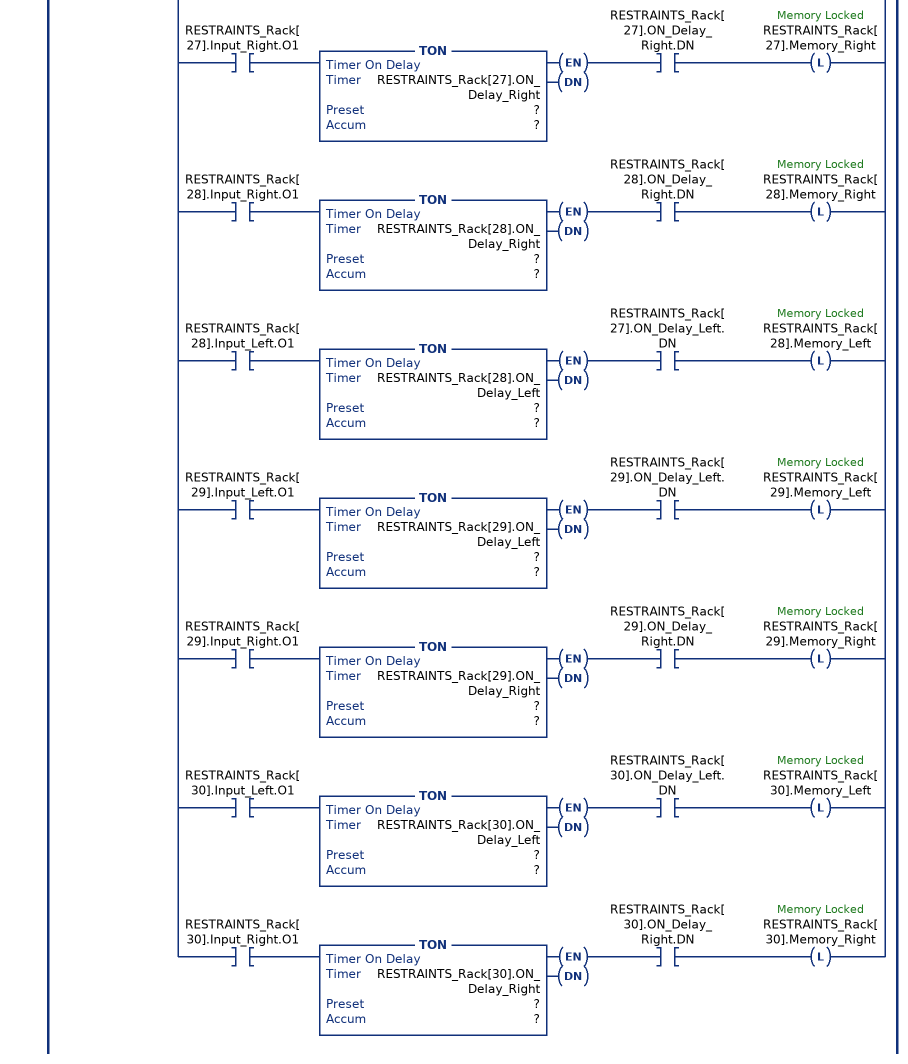
   14: XIC(Restraints_Cycle.Step_22)[XIC(RESTRAINTS_Rack[17].Input_Left.O1) TON(RESTRAINTS_Rack[17].ON_Delay_Left,?,?) XIC(RESTRAINTS_Rack[17].ON_Delay_Left.DN) OTL(RESTRAINTS_Rack[17].Memory_Left) ,XIC(RESTRAINTS_Rack[17].Input_Right.O1) TON(RESTRAINTS_Rack[17].ON_Delay_Right,?,?) XIC(RESTRAINTS_Rack[17].ON_Delay_Right.DN) OTL(RESTRAINTS_Rack[17].Memory_Right) ,XIC(RESTRAINTS_Rack[18].Input_Left.O1) TON(RESTRAINTS_Rack[18].ON_Delay_Left,?,?) XIC(RESTRAINTS_Rack[18].ON_Delay_Left.DN) OTL(RESTRAINTS_Rack[18].Memory_Left) ,XIC(RESTRAINTS_Rack[18].Input_Right.O1) TON(RESTRAINTS_Rack[18].ON_Delay_Right,?,?) XIC(RESTRAINTS_Rack[18].ON_Delay_Right.DN) OTL(RESTRAINTS_Rack[18].Memory_Right) ,XIC(RESTRAINTS_Rack[19].Input_Left.O1) TON(RESTRAINTS_Rack[19].ON_Delay_Left,?,?) XIC(RESTRAINTS_Rack[19].ON_Delay_Left.DN) OTL(RESTRAINTS_Rack[19].Memory_Left) ,XIC(RESTRAINTS_Rack[19].Input_Right.O1) TON(RESTRAINTS_Rack[19].ON_Delay_Right,?,?) XIC(RESTRAINTS_Rack[19].ON_Delay_Right.DN) OTL(RESTRAINTS_Rack[19].Memory_Right) ,XIC(RESTRAINTS_Rack[20].Input_Left.O1) TON(RESTRAINTS_Rack[20].ON_Delay_Left,?,?) XIC(RESTRAINTS_Rack[20].ON_Delay_Left.DN) OTL(RESTRAINTS_Rack[20].Memory_Left) ,XIC(RESTRAINTS_Rack[20].Input_Right.O1) TON(RESTRAINTS_Rack[20].ON_Delay_Right,?,?) XIC(RESTRAINTS_Rack[20].ON_Delay_Right.DN) OTL(RESTRAINTS_Rack[20].Memory_Right) ,XIC(RESTRAINTS_Rack[21].Input_Left.O1) TON(RESTRAINTS_Rack[21].ON_Delay_Left,?,?) XIC(RESTRAINTS_Rack[21].ON_Delay_Left.DN) OTL(RESTRAINTS_Rack[21].Memory_Left) ,XIC(RESTRAINTS_Rack[21].Input_Right.O1) TON(RESTRAINTS_Rack[21].ON_Delay_Right,?,?) XIC(RESTRAINTS_Rack[21].ON_Delay_Right.DN) OTL(RESTRAINTS_Rack[21].Memory_Right) ,XIC(RESTRAINTS_Rack[22].Input_Left.O1) TON(RESTRAINTS_Rack[22].ON_Delay_Left,?,?) XIC(RESTRAINTS_Rack[22].ON_Delay_Left.DN) OTL(RESTRAINTS_Rack[22].Memory_Left) ,XIC(RESTRAINTS_Rack[22].Input_Right.O1) TON(RESTRAINTS_Rack[22].ON_Delay_Right,?,?) XIC(RESTRAINTS_Rack[22].ON_Delay_Right.DN) OTL(RESTRAINTS_Rack[22].Memory_Right) ,XIC(RESTRAINTS_Rack[23].Input_Left.O1) TON(RESTRAINTS_Rack[23].ON_Delay_Left,?,?) XIC(RESTRAINTS_Rack[23].ON_Delay_Left.DN) OTL(RESTRAINTS_Rack[23].Memory_Left) ,XIC(RESTRAINTS_Rack[23].Input_Right.O1) TON(RESTRAINTS_Rack[23].ON_Delay_Right,?,?) XIC(RESTRAINTS_Rack[23].ON_Delay_Right.DN) OTL(RESTRAINTS_Rack[23].Memory_Right) ,XIC(RESTRAINTS_Rack[24].Input_Left.O1) TON(RESTRAINTS_Rack[24].ON_Delay_Left,?,?) XIC(RESTRAINTS_Rack[24].ON_Delay_Left.DN) OTL(RESTRAINTS_Rack[24].Memory_Left) ,XIC(RESTRAINTS_Rack[24].Input_Right.O1) TON(RESTRAINTS_Rack[24].ON_Delay_Right,?,?) XIC(RESTRAINTS_Rack[24].ON_Delay_Right.DN) OTL(RESTRAINTS_Rack[24].Memory_Right) ,XIC(RESTRAINTS_Rack[25].Input_Left.O1) TON(RESTRAINTS_Rack[25].ON_Delay_Left,?,?) XIC(RESTRAINTS_Rack[25].ON_Delay_Left.DN) OTL(RESTRAINTS_Rack[25].Memory_Left) ,XIC(RESTRAINTS_Rack[25].Input_Right.O1) TON(RESTRAINTS_Rack[25].ON_Delay_Right,?,?) XIC(RESTRAINTS_Rack[25].ON_Delay_Right.DN) OTL(RESTRAINTS_Rack[25].Memory_Right) ,XIC(RESTRAINTS_Rack[26].Input_Left.O1) TON(RESTRAINTS_Rack[26].ON_Delay_Left,?,?) XIC(RESTRAINTS_Rack[26].ON_Delay_Left.DN) OTL(RESTRAINTS_Rack[26].Memory_Left) ,XIC(RESTRAINTS_Rack[26].Input_Right.O1) TON(RESTRAINTS_Rack[26].ON_Delay_Right,?,?) XIC(RESTRAINTS_Rack[26].ON_Delay_Right.DN) OTL(RESTRAINTS_Rack[26].Memory_Right) ,XIC(RESTRAINTS_Rack[27].Input_Left.O1) TON(RESTRAINTS_Rack[27].ON_Delay_Left,?,?) XIC(RESTRAINTS_Rack[27].ON_Delay_Left.DN) OTL(RESTRAINTS_Rack[27].Memory_Left) ,XIC(RESTRAINTS_Rack[27].Input_Right.O1) TON(RESTRAINTS_Rack[27].ON_Delay_Right,?,?) XIC(RESTRAINTS_Rack[27].ON_Delay_Right.DN) OTL(RESTRAINTS_Rack[27].Memory_Right) ,XIC(RESTRAINTS_Rack[28].Input_Right.O1) TON(RESTRAINTS_Rack[28].ON_Delay_Right,?,?) XIC(RESTRAINTS_Rack[28].ON_Delay_Right.DN) OTL(RESTRAINTS_Rack[28].Memory_Right) ,XIC(RESTRAINTS_Rack[28].Input_Left.O1) TON(RESTRAINTS_Rack[28].ON_Delay_Left,?,?) XIC(RESTRAINTS_Rack[27].ON_Delay_Left.DN) OTL(RESTRAINTS_Rack[28].Memory_Left) ,XIC(RESTRAINTS_Rack[29].Input_Left.O1) TON(RESTRAINTS_Rack[29].ON_Delay_Left,?,?) XIC(RESTRAINTS_Rack[29].ON_Delay_Left.DN) OTL(RESTRAINTS_Rack[29].Memory_Left) ,XIC(RESTRAINTS_Rack[29].Input_Right.O1) TON(RESTRAINTS_Rack[29].ON_Delay_Right,?,?) XIC(RESTRAINTS_Rack[29].ON_Delay_Right.DN) OTL(RESTRAINTS_Rack[29].Memory_Right) ,XIC(RESTRAINTS_Rack[30].Input_Left.O1) TON(RESTRAINTS_Rack[30].ON_Delay_Left,?,?) XIC(RESTRAINTS_Rack[30].ON_Delay_Left.DN) OTL(RESTRAINTS_Rack[30].Memory_Left) ,XIC(RESTRAINTS_Rack[30].Input_Right.O1) TON(RESTRAINTS_Rack[30].ON_Delay_Right,?,?) XIC(RESTRAINTS_Rack[30].ON_Delay_Right.DN) OTL(RESTRAINTS_Rack[30].Memory_Right) ];
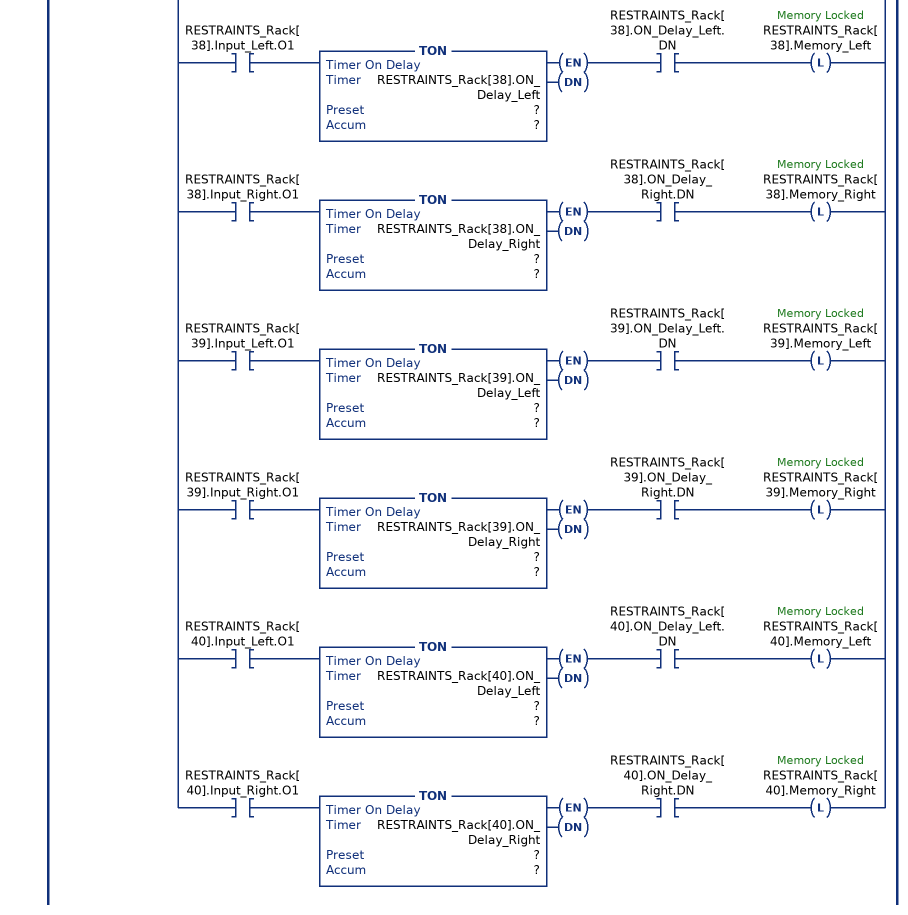
   15: XIC(Restraints_Cycle.Step_22)[XIC(RESTRAINTS_Rack[31].Input_Left.O1) TON(RESTRAINTS_Rack[31].ON_Delay_Left,?,?) XIC(RESTRAINTS_Rack[31].ON_Delay_Left.DN) OTL(RESTRAINTS_Rack[31].Memory_Left) ,XIC(RESTRAINTS_Rack[31].Input_Right.O1) TON(RESTRAINTS_Rack[31].ON_Delay_Right,?,?) XIC(RESTRAINTS_Rack[31].ON_Delay_Right.DN) OTL(RESTRAINTS_Rack[31].Memory_Right) ,XIC(RESTRAINTS_Rack[32].Input_Left.O1) TON(RESTRAINTS_Rack[32].ON_Delay_Left,?,?) XIC(RESTRAINTS_Rack[32].ON_Delay_Left.DN) OTL(RESTRAINTS_Rack[32].Memory_Left) ,XIC(RESTRAINTS_Rack[32].Input_Right.O1) TON(RESTRAINTS_Rack[32].ON_Delay_Right,?,?) XIC(RESTRAINTS_Rack[32].ON_Delay_Right.DN) OTL(RESTRAINTS_Rack[32].Memory_Right) ,XIC(RESTRAINTS_Rack[33].Input_Left.O1) TON(RESTRAINTS_Rack[33].ON_Delay_Left,?,?) XIC(RESTRAINTS_Rack[33].ON_Delay_Left.DN) OTL(RESTRAINTS_Rack[33].Memory_Left) ,XIC(RESTRAINTS_Rack[33].Input_Right.O1) TON(RESTRAINTS_Rack[33].ON_Delay_Right,?,?) XIC(RESTRAINTS_Rack[33].ON_Delay_Right.DN) OTL(RESTRAINTS_Rack[33].Memory_Right) ,XIC(RESTRAINTS_Rack[34].Input_Left.O1) TON(RESTRAINTS_Rack[34].ON_Delay_Left,?,?) XIC(RESTRAINTS_Rack[34].ON_Delay_Left.DN) OTL(RESTRAINTS_Rack[34].Memory_Left) ,XIC(RESTRAINTS_Rack[34].Input_Right.O1) TON(RESTRAINTS_Rack[34].ON_Delay_Right,?,?) XIC(RESTRAINTS_Rack[34].ON_Delay_Right.DN) OTL(RESTRAINTS_Rack[34].Memory_Right) ,XIC(RESTRAINTS_Rack[35].Input_Left.O1) TON(RESTRAINTS_Rack[35].ON_Delay_Left,?,?) XIC(RESTRAINTS_Rack[35].ON_Delay_Left.DN) OTL(RESTRAINTS_Rack[35].Memory_Left) ,XIC(RESTRAINTS_Rack[35].Input_Right.O1) TON(RESTRAINTS_Rack[35].ON_Delay_Right,?,?) XIC(RESTRAINTS_Rack[35].ON_Delay_Right.DN) OTL(RESTRAINTS_Rack[35].Memory_Right) ,XIC(RESTRAINTS_Rack[36].Input_Left.O1) TON(RESTRAINTS_Rack[36].ON_Delay_Left,?,?) XIC(RESTRAINTS_Rack[36].ON_Delay_Left.DN) OTL(RESTRAINTS_Rack[36].Memory_Left) ,XIC(RESTRAINTS_Rack[36].Input_Right.O1) TON(RESTRAINTS_Rack[36].ON_Delay_Right,?,?) XIC(RESTRAINTS_Rack[36].ON_Delay_Right.DN) OTL(RESTRAINTS_Rack[36].Memory_Right) ,XIC(RESTRAINTS_Rack[37].Input_Left.O1) TON(RESTRAINTS_Rack[37].ON_Delay_Left,?,?) XIC(RESTRAINTS_Rack[37].ON_Delay_Left.DN) OTL(RESTRAINTS_Rack[37].Memory_Left) ,XIC(RESTRAINTS_Rack[37].Input_Right.O1) TON(RESTRAINTS_Rack[37].ON_Delay_Right,?,?) XIC(RESTRAINTS_Rack[37].ON_Delay_Right.DN) OTL(RESTRAINTS_Rack[37].Memory_Right) ,XIC(RESTRAINTS_Rack[38].Input_Left.O1) TON(RESTRAINTS_Rack[38].ON_Delay_Left,?,?) XIC(RESTRAINTS_Rack[38].ON_Delay_Left.DN) OTL(RESTRAINTS_Rack[38].Memory_Left) ,XIC(RESTRAINTS_Rack[38].Input_Right.O1) TON(RESTRAINTS_Rack[38].ON_Delay_Right,?,?) XIC(RESTRAINTS_Rack[38].ON_Delay_Right.DN) OTL(RESTRAINTS_Rack[38].Memory_Right) ,XIC(RESTRAINTS_Rack[39].Input_Left.O1) TON(RESTRAINTS_Rack[39].ON_Delay_Left,?,?) XIC(RESTRAINTS_Rack[39].ON_Delay_Left.DN) OTL(RESTRAINTS_Rack[39].Memory_Left) ,XIC(RESTRAINTS_Rack[39].Input_Right.O1) TON(RESTRAINTS_Rack[39].ON_Delay_Right,?,?) XIC(RESTRAINTS_Rack[39].ON_Delay_Right.DN) OTL(RESTRAINTS_Rack[39].Memory_Right) ,XIC(RESTRAINTS_Rack[40].Input_Left.O1) TON(RESTRAINTS_Rack[40].ON_Delay_Left,?,?) XIC(RESTRAINTS_Rack[40].ON_Delay_Left.DN) OTL(RESTRAINTS_Rack[40].Memory_Left) ,XIC(RESTRAINTS_Rack[40].Input_Right.O1) TON(RESTRAINTS_Rack[40].ON_Delay_Right,?,?) XIC(RESTRAINTS_Rack[40].ON_Delay_Right.DN) OTL(RESTRAINTS_Rack[40].Memory_Right) ];
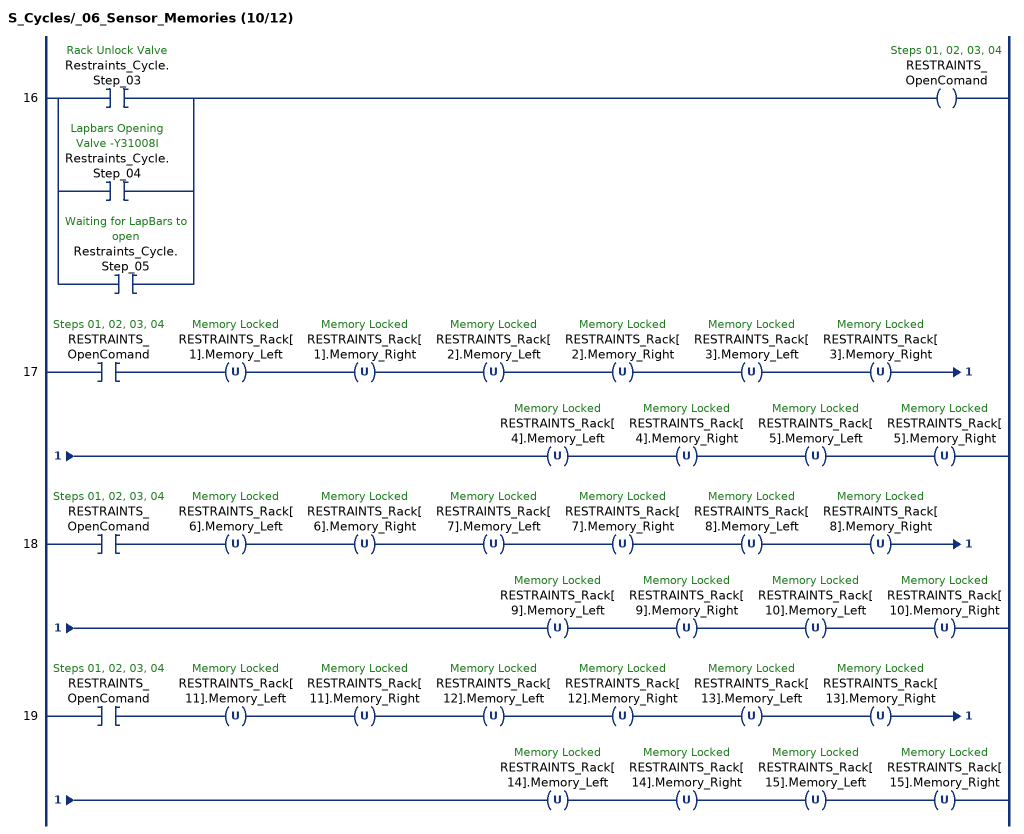
   16: [XIC(Restraints_Cycle.Step_03) ,XIC(Restraints_Cycle.Step_04) ,XIC(Restraints_Cycle.Step_05) ]OTE(RESTRAINTS_OpenComand);
   17: XIC(RESTRAINTS_OpenComand)OTU(RESTRAINTS_Rack[1].Memory_Left)OTU(RESTRAINTS_Rack[1].Memory_Right)OTU(RESTRAINTS_Rack[2].Memory_Left)OTU(RESTRAINTS_Rack[2].Memory_Right)OTU(RESTRAINTS_Rack[3].Memory_Left)OTU(RESTRAINTS_Rack[3].Memory_Right)OTU(RESTRAINTS_Rack[4].Memory_Left)OTU(RESTRAINTS_Rack[4].Memory_Right)OTU(RESTRAINTS_Rack[5].Memory_Left)OTU(RESTRAINTS_Rack[5].Memory_Right);
   18: XIC(RESTRAINTS_OpenComand)OTU(RESTRAINTS_Rack[6].Memory_Left)OTU(RESTRAINTS_Rack[6].Memory_Right)OTU(RESTRAINTS_Rack[7].Memory_Left)OTU(RESTRAINTS_Rack[7].Memory_Right)OTU(RESTRAINTS_Rack[8].Memory_Left)OTU(RESTRAINTS_Rack[8].Memory_Right)OTU(RESTRAINTS_Rack[9].Memory_Left)OTU(RESTRAINTS_Rack[9].Memory_Right)OTU(RESTRAINTS_Rack[10].Memory_Left)OTU(RESTRAINTS_Rack[10].Memory_Right);
   19: XIC(RESTRAINTS_OpenComand)OTU(RESTRAINTS_Rack[11].Memory_Left)OTU(RESTRAINTS_Rack[11].Memory_Right)OTU(RESTRAINTS_Rack[12].Memory_Left)OTU(RESTRAINTS_Rack[12].Memory_Right)OTU(RESTRAINTS_Rack[13].Memory_Left)OTU(RESTRAINTS_Rack[13].Memory_Right)OTU(RESTRAINTS_Rack[14].Memory_Left)OTU(RESTRAINTS_Rack[14].Memory_Right)OTU(RESTRAINTS_Rack[15].Memory_Left)OTU(RESTRAINTS_Rack[15].Memory_Right);
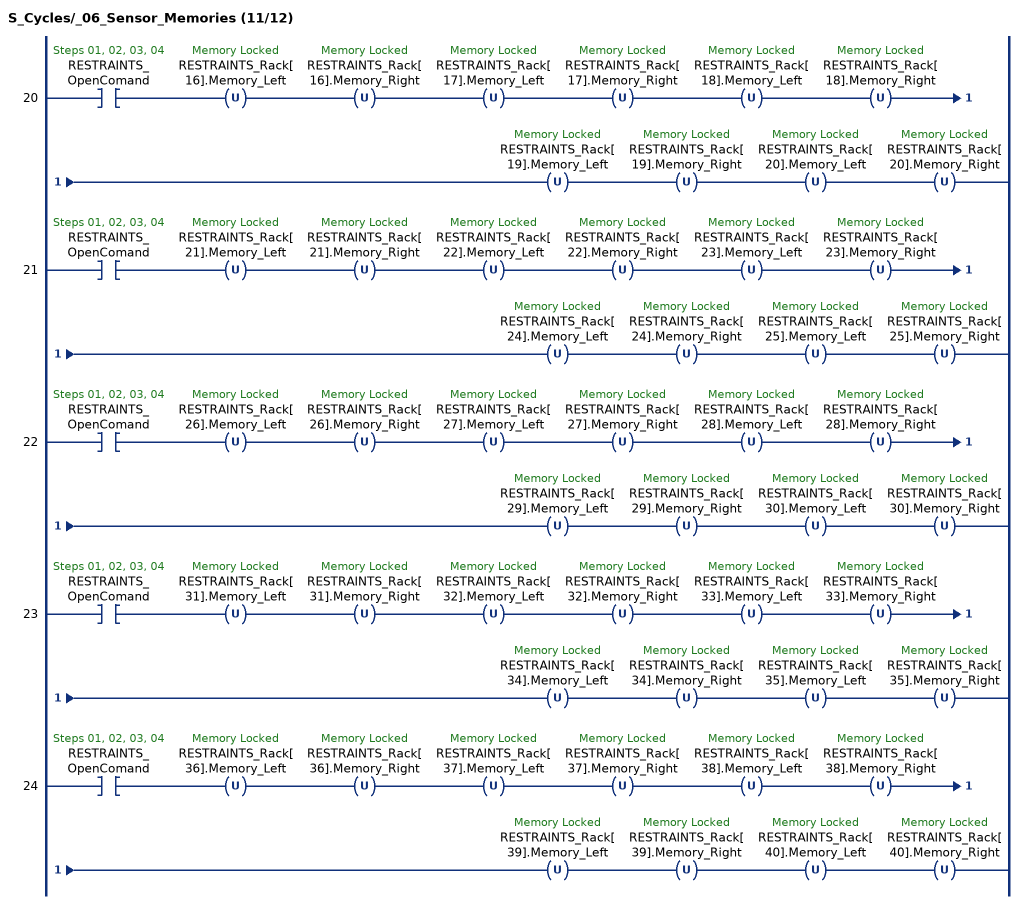
   20: XIC(RESTRAINTS_OpenComand)OTU(RESTRAINTS_Rack[16].Memory_Left)OTU(RESTRAINTS_Rack[16].Memory_Right)OTU(RESTRAINTS_Rack[17].Memory_Left)OTU(RESTRAINTS_Rack[17].Memory_Right)OTU(RESTRAINTS_Rack[18].Memory_Left)OTU(RESTRAINTS_Rack[18].Memory_Right)OTU(RESTRAINTS_Rack[19].Memory_Left)OTU(RESTRAINTS_Rack[19].Memory_Right)OTU(RESTRAINTS_Rack[20].Memory_Left)OTU(RESTRAINTS_Rack[20].Memory_Right);
   21: XIC(RESTRAINTS_OpenComand)OTU(RESTRAINTS_Rack[21].Memory_Left)OTU(RESTRAINTS_Rack[21].Memory_Right)OTU(RESTRAINTS_Rack[22].Memory_Left)OTU(RESTRAINTS_Rack[22].Memory_Right)OTU(RESTRAINTS_Rack[23].Memory_Left)OTU(RESTRAINTS_Rack[23].Memory_Right)OTU(RESTRAINTS_Rack[24].Memory_Left)OTU(RESTRAINTS_Rack[24].Memory_Right)OTU(RESTRAINTS_Rack[25].Memory_Left)OTU(RESTRAINTS_Rack[25].Memory_Right);
   22: XIC(RESTRAINTS_OpenComand)OTU(RESTRAINTS_Rack[26].Memory_Left)OTU(RESTRAINTS_Rack[26].Memory_Right)OTU(RESTRAINTS_Rack[27].Memory_Left)OTU(RESTRAINTS_Rack[27].Memory_Right)OTU(RESTRAINTS_Rack[28].Memory_Left)OTU(RESTRAINTS_Rack[28].Memory_Right)OTU(RESTRAINTS_Rack[29].Memory_Left)OTU(RESTRAINTS_Rack[29].Memory_Right)OTU(RESTRAINTS_Rack[30].Memory_Left)OTU(RESTRAINTS_Rack[30].Memory_Right);
   23: XIC(RESTRAINTS_OpenComand)OTU(RESTRAINTS_Rack[31].Memory_Left)OTU(RESTRAINTS_Rack[31].Memory_Right)OTU(RESTRAINTS_Rack[32].Memory_Left)OTU(RESTRAINTS_Rack[32].Memory_Right)OTU(RESTRAINTS_Rack[33].Memory_Left)OTU(RESTRAINTS_Rack[33].Memory_Right)OTU(RESTRAINTS_Rack[34].Memory_Left)OTU(RESTRAINTS_Rack[34].Memory_Right)OTU(RESTRAINTS_Rack[35].Memory_Left)OTU(RESTRAINTS_Rack[35].Memory_Right);
   24: XIC(RESTRAINTS_OpenComand)OTU(RESTRAINTS_Rack[36].Memory_Left)OTU(RESTRAINTS_Rack[36].Memory_Right)OTU(RESTRAINTS_Rack[37].Memory_Left)OTU(RESTRAINTS_Rack[37].Memory_Right)OTU(RESTRAINTS_Rack[38].Memory_Left)OTU(RESTRAINTS_Rack[38].Memory_Right)OTU(RESTRAINTS_Rack[39].Memory_Left)OTU(RESTRAINTS_Rack[39].Memory_Right)OTU(RESTRAINTS_Rack[40].Memory_Left)OTU(RESTRAINTS_Rack[40].Memory_Right);
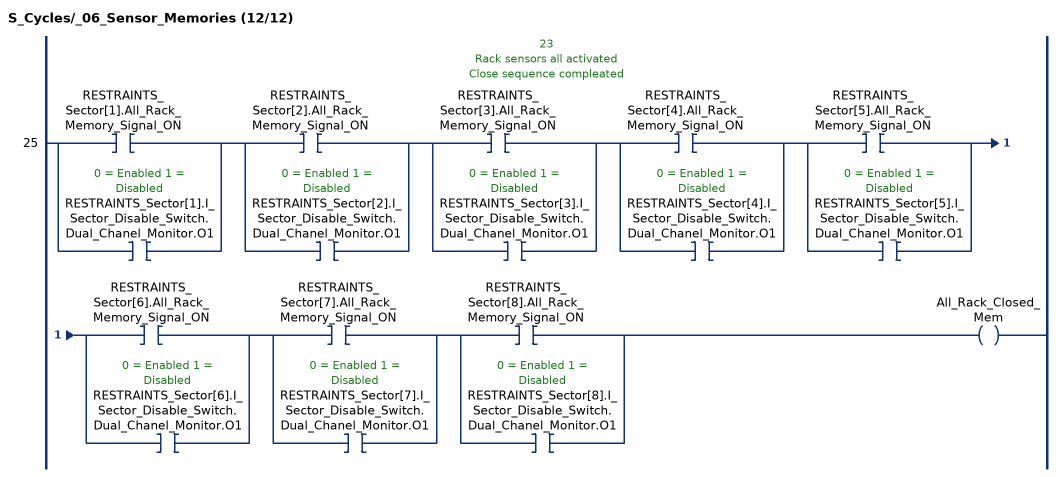
   // 23
   // Rack sensors all activated
   // Close sequence compleated
   25: [XIC(RESTRAINTS_Sector[1].All_Rack_Memory_Signal_ON) ,XIC(RESTRAINTS_Sector[1].I_Sector_Disable_Switch.Dual_Chanel_Monitor.O1) ][XIC(RESTRAINTS_Sector[2].All_Rack_Memory_Signal_ON) ,XIC(RESTRAINTS_Sector[2].I_Sector_Disable_Switch.Dual_Chanel_Monitor.O1) ][XIC(RESTRAINTS_Sector[3].All_Rack_Memory_Signal_ON) ,XIC(RESTRAINTS_Sector[3].I_Sector_Disable_Switch.Dual_Chanel_Monitor.O1) ][XIC(RESTRAINTS_Sector[4].All_Rack_Memory_Signal_ON) ,XIC(RESTRAINTS_Sector[4].I_Sector_Disable_Switch.Dual_Chanel_Monitor.O1) ][XIC(RESTRAINTS_Sector[5].All_Rack_Memory_Signal_ON) ,XIC(RESTRAINTS_Sector[5].I_Sector_Disable_Switch.Dual_Chanel_Monitor.O1) ][XIC(RESTRAINTS_Sector[6].All_Rack_Memory_Signal_ON) ,XIC(RESTRAINTS_Sector[6].I_Sector_Disable_Switch.Dual_Chanel_Monitor.O1) ][XIC(RESTRAINTS_Sector[7].All_Rack_Memory_Signal_ON) ,XIC(RESTRAINTS_Sector[7].I_Sector_Disable_Switch.Dual_Chanel_Monitor.O1) ][XIC(RESTRAINTS_Sector[8].All_Rack_Memory_Signal_ON) ,XIC(RESTRAINTS_Sector[8].I_Sector_Disable_Switch.Dual_Chanel_Monitor.O1) ]OTE(All_Rack_Closed_Mem);
END_ROUTINE

ROUTINE _99_Commands   (* ladder *)
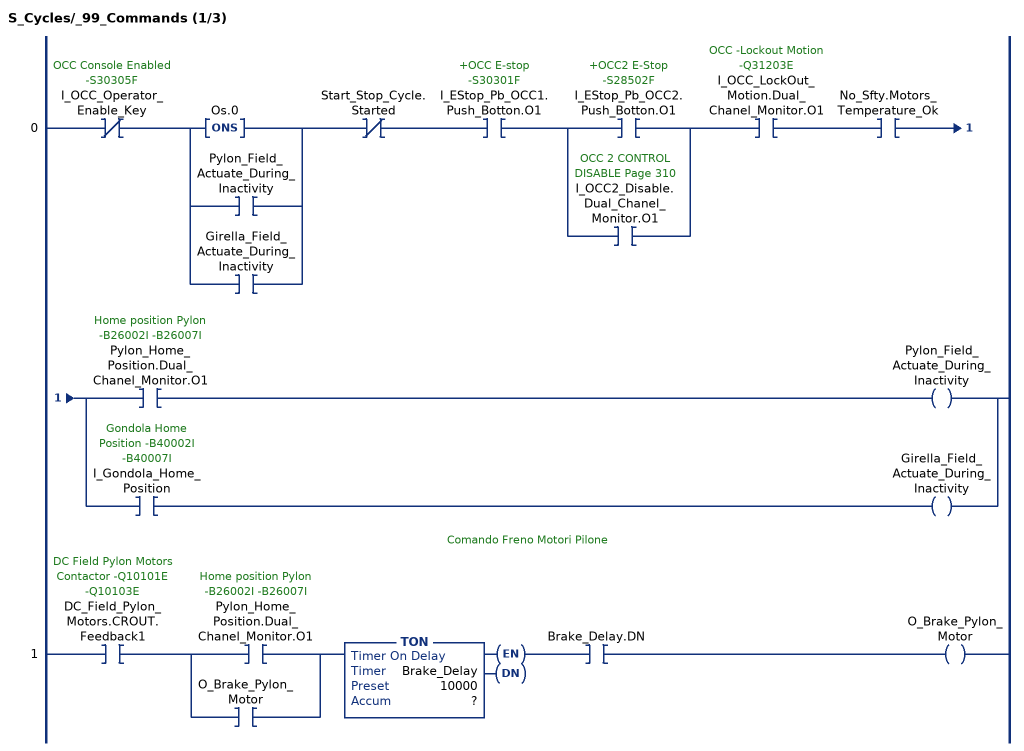
   0: XIO(I_OCC_Operator_Enable_Key)[ONS(Os.0) ,XIC(Pylon_Field_Actuate_During_Inactivity) ,XIC(Girella_Field_Actuate_During_Inactivity) ]XIO(Start_Stop_Cycle.Started)XIC(I_EStop_Pb_OCC1.Push_Botton.O1)[XIC(I_EStop_Pb_OCC2.Push_Botton.O1) ,XIC(I_OCC2_Disable.Dual_Chanel_Monitor.O1) ]XIC(I_OCC_LockOut_Motion.Dual_Chanel_Monitor.O1)XIC(No_Sfty.Motors_Temperature_Ok)[XIC(Pylon_Home_Position.Dual_Chanel_Monitor.O1) OTE(Pylon_Field_Actuate_During_Inactivity) ,XIC(I_Gondola_Home_Position) OTE(Girella_Field_Actuate_During_Inactivity) ];
   // Comando Freno Motori Pilone
   1: XIC(DC_Field_Pylon_Motors.CROUT.Feedback1)[XIC(Pylon_Home_Position.Dual_Chanel_Monitor.O1) ,XIC(O_Brake_Pylon_Motor) ]TON(Brake_Delay,?,?)XIC(Brake_Delay.DN)OTE(O_Brake_Pylon_Motor);
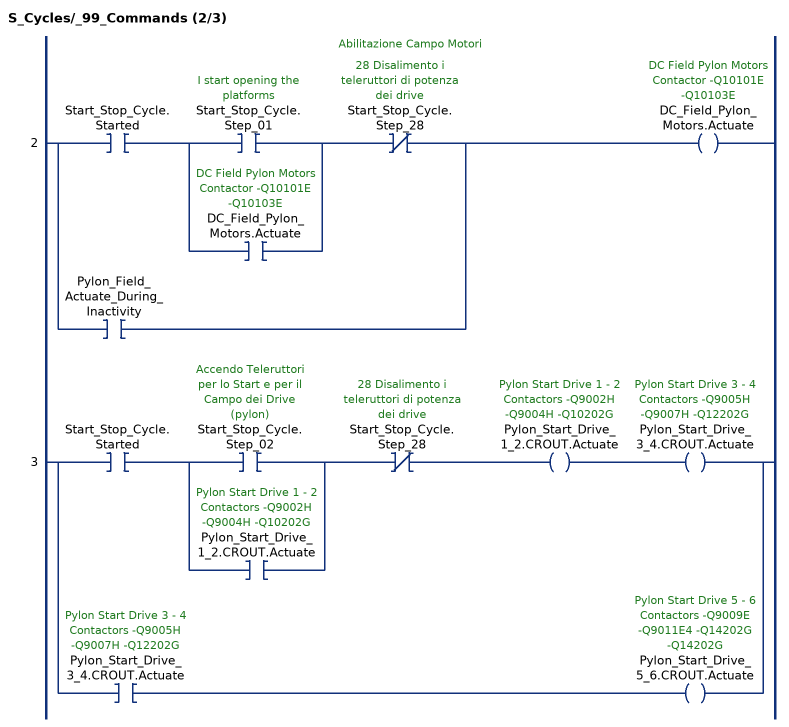
   // Abilitazione Campo Motori
   2: [XIC(Start_Stop_Cycle.Started) [XIC(Start_Stop_Cycle.Step_01) ,XIC(DC_Field_Pylon_Motors.Actuate) ] XIO(Start_Stop_Cycle.Step_28) ,XIC(Pylon_Field_Actuate_During_Inactivity) ]OTE(DC_Field_Pylon_Motors.Actuate);
   3: [XIC(Start_Stop_Cycle.Started) [XIC(Start_Stop_Cycle.Step_02) ,XIC(Pylon_Start_Drive_1_2.CROUT.Actuate) ] XIO(Start_Stop_Cycle.Step_28) OTE(Pylon_Start_Drive_1_2.CROUT.Actuate) OTE(Pylon_Start_Drive_3_4.CROUT.Actuate) ,XIC(Pylon_Start_Drive_3_4.CROUT.Actuate) OTE(Pylon_Start_Drive_5_6.CROUT.Actuate) ];
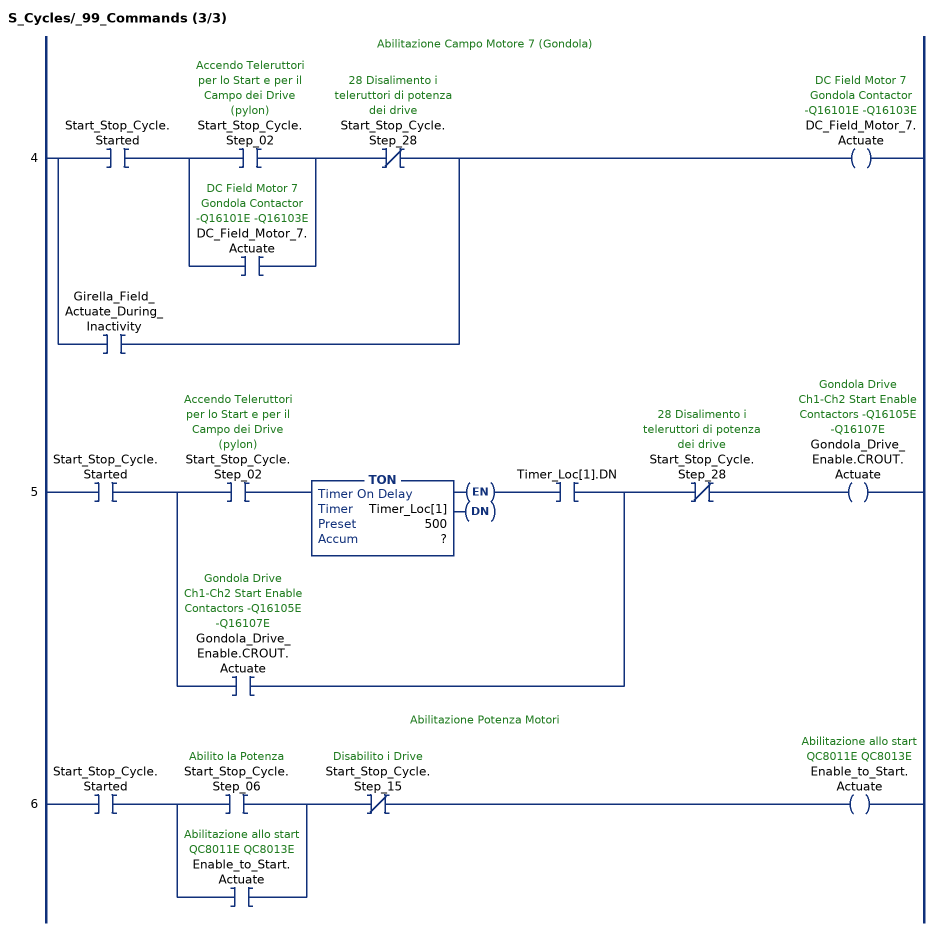
   // Abilitazione Campo Motore 7 (Gondola)
   4: [XIC(Start_Stop_Cycle.Started) [XIC(Start_Stop_Cycle.Step_02) ,XIC(DC_Field_Motor_7.Actuate) ] XIO(Start_Stop_Cycle.Step_28) ,XIC(Girella_Field_Actuate_During_Inactivity) ]OTE(DC_Field_Motor_7.Actuate);
   5: XIC(Start_Stop_Cycle.Started)[XIC(Start_Stop_Cycle.Step_02) TON(Timer_Loc[1],?,?) XIC(Timer_Loc[1].DN) ,XIC(Gondola_Drive_Enable.CROUT.Actuate) ]XIO(Start_Stop_Cycle.Step_28)OTE(Gondola_Drive_Enable.CROUT.Actuate);
   // Abilitazione Potenza Motori
   6: XIC(Start_Stop_Cycle.Started)[XIC(Start_Stop_Cycle.Step_06) ,XIC(Enable_to_Start.Actuate) ]XIO(Start_Stop_Cycle.Step_15)OTE(Enable_to_Start.Actuate);
END_ROUTINE

ROUTINE Main   (* ladder *)
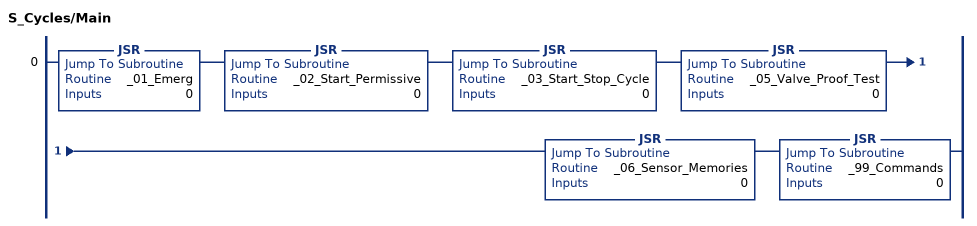
   0: JSR(_01_Emerg,0)JSR(_02_Start_Permissive,0)JSR(_03_Start_Stop_Cycle,0)JSR(_05_Valve_Proof_Test,0)JSR(_06_Sensor_Memories,0)JSR(_99_Commands,0);
END_ROUTINE
END_PROGRAM
